// TIA Portal project "XSFW_TIA32801_A0" (V15.1) (continued)
REGION Network 14: Agrupa las fallas del proceso en una marca
   RUNG wire#powerrail
      I_Contact( "Fallas"."area de recorrido libre del pusher" )
      I_Contact( "Fallas"."caja trabada a la salida" )
      I_Contact( "Fallas".emergencia )
      I_Contact( "Fallas"."Falla de programación concatenadoras 1" )
      I_Contact( "Fallas"."Falla de programación concatenadoras 2" )
      I_Contact( "Fallas"."Falla de programación prioritarias 1" )
      I_Contact( "Fallas"."Falla de programación prioritarias 2" )
      I_Contact( "Fallas"."Falla en rele cadena" )
      I_Contact( "Fallas"."Falla en sensor de encolado" )
      I_Contact( "Fallas".falla_encoder )
      I_Contact( "Fallas".falla_sns_bsucc_ab )
      I_Contact( "Fallas".falla_sns_bsucc_ar )
      I_Contact( "Fallas"."Incrongruencia pusher" )
      I_Contact( "Fallas"."proteccion de torque" )
      I_Contact( "Fallas"."Falla en sensores del Pusher" )
      I_Contact( "Fallas"."Sensor pusher hacia adelante" )
      I_Contact( "Fallas"."Sin pegamento en el depósito" )
      I_Contact( "Fallas"."Falla de caja cerrada en cadena" )
      Coil( "Serie de fallas" )
   END_RUNG
   // the same network as SCL:
   "Serie de fallas" := NOT "Fallas"."area de recorrido libre del pusher" AND NOT "Fallas"."caja trabada a la salida" AND NOT "Fallas".emergencia AND NOT "Fallas"."Falla de programación concatenadoras 1" AND NOT "Fallas"."Falla de programación concatenadoras 2" AND NOT "Fallas"."Falla de programación prioritarias 1" AND NOT "Fallas"."Falla de programación prioritarias 2" AND NOT "Fallas"."Falla en rele cadena" AND NOT "Fallas"."Falla en sensor de encolado" AND NOT "Fallas".falla_encoder AND NOT "Fallas".falla_sns_bsucc_ab AND NOT "Fallas".falla_sns_bsucc_ar AND NOT "Fallas"."Incrongruencia pusher" AND NOT "Fallas"."proteccion de torque" AND NOT "Fallas"."Falla en sensores del Pusher" AND NOT "Fallas"."Sensor pusher hacia adelante" AND NOT "Fallas"."Sin pegamento en el depósito" AND NOT "Fallas"."Falla de caja cerrada en cadena";
END_REGION

REGION Network 15: Fallas en sensor atras del Pusher
   "Timer_DB7".TON(IN := "1s8" AND "oM_pusher" AND NOT "iSNSpush_atras", PT := T#350MS);
   "Fallas"."Falla en sensores del Pusher" := "Timer_DB7".Q;
END_REGION

REGION Network 16: Fallas en sensor adelante del Pusher
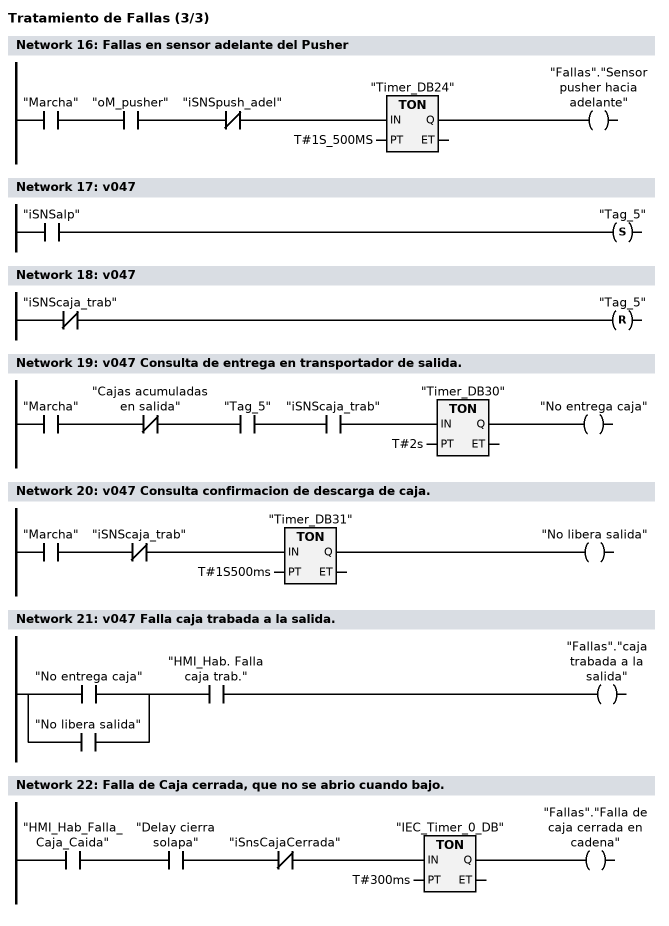
   "Timer_DB24".TON(IN := "Marcha" AND "oM_pusher" AND NOT "iSNSpush_adel", PT := T#1S_500MS);
   "Fallas"."Sensor pusher hacia adelante" := "Timer_DB24".Q;
END_REGION

REGION Network 17: v047
   RUNG wire#powerrail
      Contact( "iSNSalp" )
      S_Coil( "Tag_5" )
   END_RUNG
   // the same network as SCL:
   IF "iSNSalp" THEN "Tag_5" := TRUE; END_IF;
END_REGION

REGION Network 18: v047
   RUNG wire#powerrail
      I_Contact( "iSNScaja_trab" )
      R_Coil( "Tag_5" )
   END_RUNG
   // the same network as SCL:
   IF NOT "iSNScaja_trab" THEN "Tag_5" := FALSE; END_IF;
END_REGION

REGION Network 19: v047 Consulta de entrega en transportador de salida.
   "Timer_DB30".TON(IN := "Marcha" AND NOT "Cajas acumuladas en salida" AND "Tag_5" AND "iSNScaja_trab",
                    PT := T#2s);
   "No entrega caja" := "Timer_DB30".Q;
END_REGION

REGION Network 20: v047 Consulta confirmacion de descarga de caja.
   "Timer_DB31".TON(IN := "Marcha" AND NOT "iSNScaja_trab", PT := T#1S500ms);
   "No libera salida" := "Timer_DB31".Q;
END_REGION

REGION Network 21: v047 Falla caja trabada a la salida.
   RUNG wire#powerrail
      Contact( "No entrega caja" )
      wire#w1
      Contact( "HMI_Hab. Falla caja trab." )
      Coil( "Fallas"."caja trabada a la salida" )
   END_RUNG
   RUNG wire#powerrail
      Contact( "No libera salida" )
   END_RUNG wire#w1
   // the same network as SCL:
   "Fallas"."caja trabada a la salida" := ("No entrega caja" OR "No libera salida") AND "HMI_Hab. Falla caja trab.";
END_REGION

REGION Network 22: Falla de Caja cerrada, que no se abrio cuando bajo.
   "IEC_Timer_0_DB".TON(IN := "HMI_Hab_Falla_Caja_Caida" AND "Delay cierra solapa" AND NOT "iSnsCajaCerrada",
                        PT := T#300ms);
   "Fallas"."Falla de caja cerrada en cadena" := "IEC_Timer_0_DB".Q;
END_REGION
END_FUNCTION

FUNCTION "Salidas" : Void   // FC17, LAD
TITLE = Salidas del proceso (Modo Automático y Manual)
{ S7_Optimized_Access := 'TRUE' }
VERSION : 0.1
   VAR_TEMP   // added for the SCL form of the ladder/FBD networks
      _w1 : Bool;
   END_VAR
BEGIN

REGION Network 1: Activa la línea de emergencia del PLC
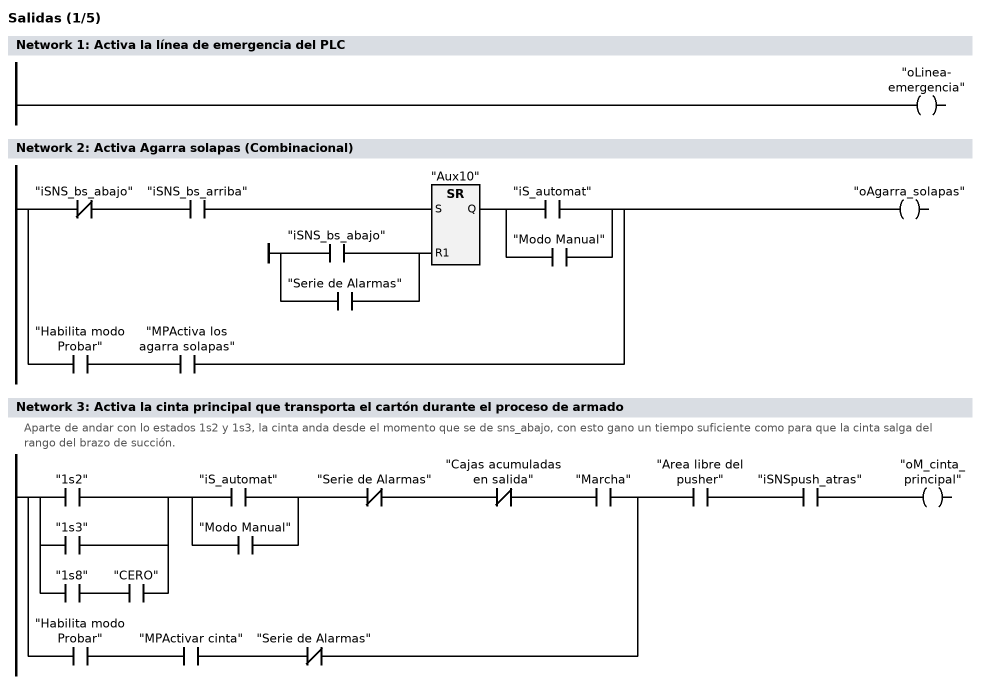
   RUNG wire#powerrail
      Coil( "oLinea-emergencia" )
   END_RUNG
   // the same network as SCL:
   "oLinea-emergencia" := TRUE;
END_REGION

REGION Network 2: Activa Agarra solapas (Combinacional)
   RUNG wire#powerrail
      I_Contact( "iSNS_bs_abajo" )
      Contact( "iSNS_bs_arriba" )
      S_SR(operand := "Aux10", r1 := wire#w1)
      wire#w2
      Contact( "iS_automat" )
      wire#w3
      Coil( "oAgarra_solapas" )
   END_RUNG
   RUNG wire#powerrail
      Contact( "iSNS_bs_abajo" )
   END_RUNG wire#w1
   RUNG wire#powerrail
      Contact( "Serie de Alarmas" )
   END_RUNG wire#w1
   RUNG wire#w2
      Contact( "Modo Manual" )
   END_RUNG wire#w3
   RUNG wire#powerrail
      Contact( "Habilita modo Probar" )
      Contact( "MPActiva los agarra solapas" )
   END_RUNG wire#w3
   // the same network as SCL:
   IF NOT "iSNS_bs_abajo" AND "iSNS_bs_arriba" THEN
       "Aux10" := TRUE;   // SR flip-flop
   END_IF;
   IF "iSNS_bs_abajo" OR "Serie de Alarmas" THEN "Aux10" := FALSE; END_IF;
   "oAgarra_solapas" := ("Aux10" AND ("iS_automat" OR "Modo Manual")) OR ("Habilita modo Probar" AND "MPActiva los agarra solapas");
END_REGION

REGION Network 3: Activa la cinta principal que transporta el cartón durante el proceso de armado
   // Aparte de andar con lo estados 1s2 y 1s3, la cinta anda desde el momento que se de sns_abajo, con esto gano un tiempo suficiente como para que la cinta salga del rango del brazo de succión.
   RUNG wire#powerrail
      Contact( "1s2" )
      wire#w1
      Contact( "iS_automat" )
      wire#w2
      I_Contact( "Serie de Alarmas" )
      I_Contact( "Cajas acumuladas en salida" )
      Contact( "Marcha" )
      wire#w3
      Contact( "Area libre del pusher" )
      Contact( "iSNSpush_atras" )
      Coil( "oM_cinta_principal" )
   END_RUNG
   RUNG wire#powerrail
      Contact( "1s3" )
   END_RUNG wire#w1
   RUNG wire#powerrail
      Contact( "1s8" )
      Contact( "CERO" )
   END_RUNG wire#w1
   RUNG wire#w1
      Contact( "Modo Manual" )
   END_RUNG wire#w2
   RUNG wire#powerrail
      Contact( "Habilita modo Probar" )
      Contact( "MPActivar cinta" )
      I_Contact( "Serie de Alarmas" )
   END_RUNG wire#w3
   // the same network as SCL:
   "oM_cinta_principal" := ((("1s2" OR "1s3" OR ("1s8" AND "CERO")) AND ("iS_automat" OR "Modo Manual") AND NOT "Serie de Alarmas" AND NOT "Cajas acumuladas en salida" AND "Marcha") OR ("Habilita modo Probar" AND "MPActivar cinta" AND NOT "Serie de Alarmas")) AND "Area libre del pusher" AND "iSNSpush_atras";
END_REGION

REGION Network 4: Activa la boquilla encoladora.
   // Activa la boquilla encoladora a partir de determinados valores del encoder.El sensor de área de encolado se utiliza para fines de seguridad. El inicio de encolado se valida con la marca "aux encol 2"
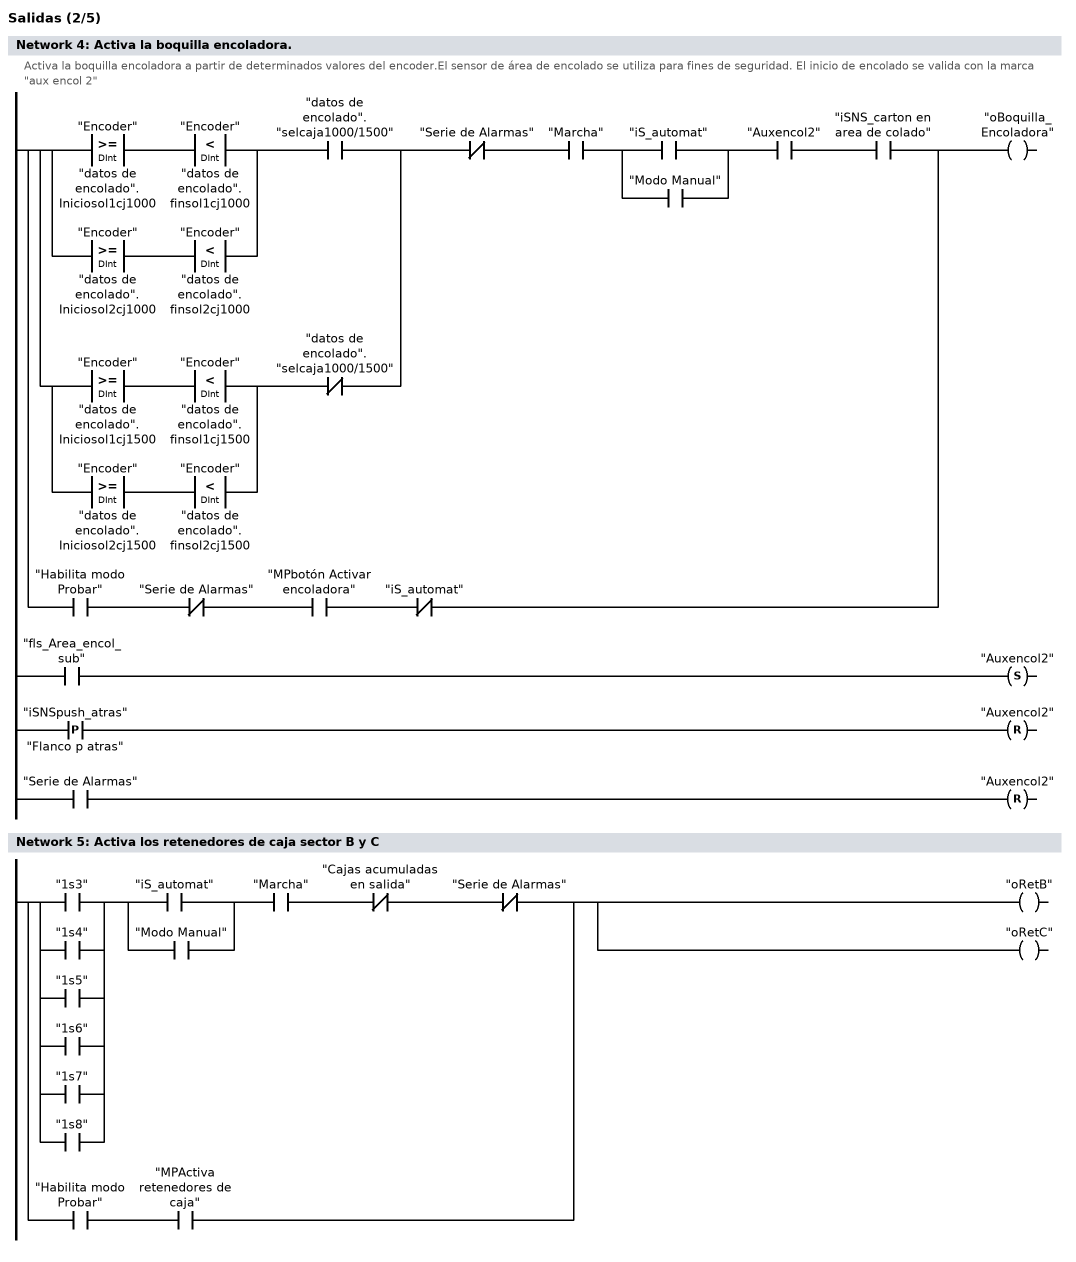
   RUNG wire#powerrail
      { S7_Templates := "SrcType := DInt" } GE_Contact(in1 := "Encoder", in2 := "datos de encolado".Iniciosol1cj1000)
      { S7_Templates := "SrcType := DInt" } LT_Contact(in1 := "Encoder", in2 := "datos de encolado".finsol1cj1000)
      wire#w1
      Contact( "datos de encolado"."selcaja1000/1500" )
      wire#w2
      I_Contact( "Serie de Alarmas" )
      Contact( "Marcha" )
      wire#w4
      Contact( "iS_automat" )
      wire#w5
      Contact( "Auxencol2" )
      Contact( "iSNS_carton en area de colado" )
      wire#w6
      Coil( "oBoquilla_Encoladora" )
   END_RUNG
   RUNG wire#powerrail
      { S7_Templates := "SrcType := DInt" } GE_Contact(in1 := "Encoder", in2 := "datos de encolado".Iniciosol2cj1000)
      { S7_Templates := "SrcType := DInt" } LT_Contact(in1 := "Encoder", in2 := "datos de encolado".finsol2cj1000)
   END_RUNG wire#w1
   RUNG wire#powerrail
      { S7_Templates := "SrcType := DInt" } GE_Contact(in1 := "Encoder", in2 := "datos de encolado".Iniciosol1cj1500)
      { S7_Templates := "SrcType := DInt" } LT_Contact(in1 := "Encoder", in2 := "datos de encolado".finsol1cj1500)
      wire#w3
      I_Contact( "datos de encolado"."selcaja1000/1500" )
   END_RUNG wire#w2
   RUNG wire#powerrail
      { S7_Templates := "SrcType := DInt" } GE_Contact(in1 := "Encoder", in2 := "datos de encolado".Iniciosol2cj1500)
      { S7_Templates := "SrcType := DInt" } LT_Contact(in1 := "Encoder", in2 := "datos de encolado".finsol2cj1500)
   END_RUNG wire#w3
   RUNG wire#w4
      Contact( "Modo Manual" )
   END_RUNG wire#w5
   RUNG wire#powerrail
      Contact( "Habilita modo Probar" )
      I_Contact( "Serie de Alarmas" )
      Contact( "MPbotón Activar encoladora" )
      I_Contact( "iS_automat" )
   END_RUNG wire#w6
   RUNG wire#powerrail
      Contact( "fls_Area_encol_sub" )
      S_Coil( "Auxencol2" )
   END_RUNG
   RUNG wire#powerrail
      P_Contact(operand := "iSNSpush_atras", bit := "Flanco p atras")
      R_Coil( "Auxencol2" )
   END_RUNG
   RUNG wire#powerrail
      Contact( "Serie de Alarmas" )
      R_Coil( "Auxencol2" )
   END_RUNG
   // the same network as SCL:
   "oBoquilla_Encoladora" := (((((("Encoder" >= "datos de encolado".Iniciosol1cj1000) AND ("Encoder" < "datos de encolado".finsol1cj1000)) OR (("Encoder" >= "datos de encolado".Iniciosol2cj1000) AND ("Encoder" < "datos de encolado".finsol2cj1000))) AND "datos de encolado"."selcaja1000/1500") OR (((("Encoder" >= "datos de encolado".Iniciosol1cj1500) AND ("Encoder" < "datos de encolado".finsol1cj1500)) OR (("Encoder" >= "datos de encolado".Iniciosol2cj1500) AND ("Encoder" < "datos de encolado".finsol2cj1500))) AND NOT "datos de encolado"."selcaja1000/1500")) AND NOT "Serie de Alarmas" AND "Marcha" AND ("iS_automat" OR "Modo Manual") AND "Auxencol2" AND "iSNS_carton en area de colado") OR ("Habilita modo Probar" AND NOT "Serie de Alarmas" AND "MPbotón Activar encoladora" AND NOT "iS_automat");
   IF "fls_Area_encol_sub" THEN "Auxencol2" := TRUE; END_IF;
   #_w1 := "iSNSpush_atras" AND NOT "Flanco p atras";   // rising edge of "iSNSpush_atras"
   "Flanco p atras" := "iSNSpush_atras";
   IF #_w1 THEN "Auxencol2" := FALSE; END_IF;
   IF "Serie de Alarmas" THEN "Auxencol2" := FALSE; END_IF;
END_REGION

REGION Network 5: Activa los retenedores de caja sector B y C
   RUNG wire#powerrail
      Contact( "1s3" )
      wire#w1
      Contact( "iS_automat" )
      wire#w2
      Contact( "Marcha" )
      I_Contact( "Cajas acumuladas en salida" )
      I_Contact( "Serie de Alarmas" )
      wire#w3
      Coil( "oRetB" )
   END_RUNG
   RUNG wire#powerrail
      Contact( "1s4" )
   END_RUNG wire#w1
   RUNG wire#powerrail
      Contact( "1s5" )
   END_RUNG wire#w1
   RUNG wire#powerrail
      Contact( "1s6" )
   END_RUNG wire#w1
   RUNG wire#powerrail
      Contact( "1s7" )
   END_RUNG wire#w1
   RUNG wire#powerrail
      Contact( "1s8" )
   END_RUNG wire#w1
   RUNG wire#w1
      Contact( "Modo Manual" )
   END_RUNG wire#w2
   RUNG wire#powerrail
      Contact( "Habilita modo Probar" )
      Contact( "MPActiva retenedores de caja" )
   END_RUNG wire#w3
   RUNG wire#w3
      Coil( "oRetC" )
   END_RUNG
   // the same network as SCL:
   "oRetB" := (("1s3" OR "1s4" OR "1s5" OR "1s6" OR "1s7" OR "1s8") AND ("iS_automat" OR "Modo Manual") AND "Marcha" AND NOT "Cajas acumuladas en salida" AND NOT "Serie de Alarmas") OR ("Habilita modo Probar" AND "MPActiva retenedores de caja");
   "oRetC" := "oRetB";
END_REGION

REGION Network 6
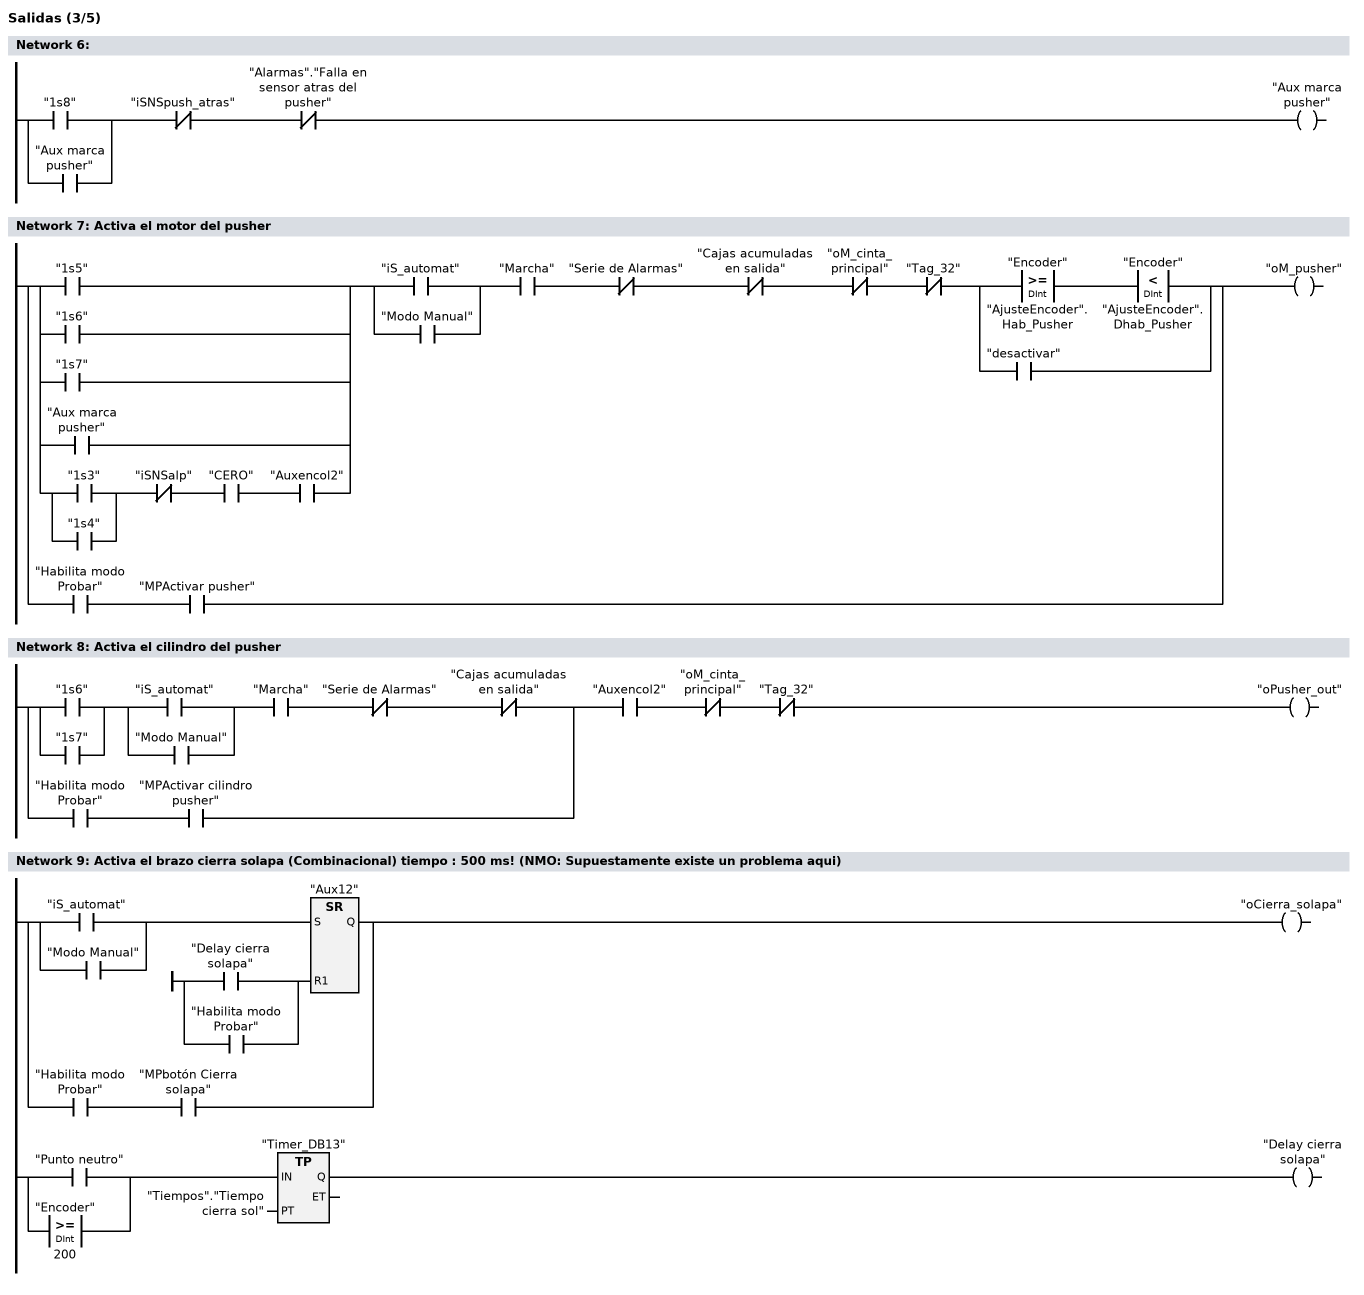
   RUNG wire#powerrail
      Contact( "1s8" )
      wire#w1
      I_Contact( "iSNSpush_atras" )
      I_Contact( "Alarmas"."Falla en sensor atras del pusher" )
      Coil( "Aux marca pusher" )
   END_RUNG
   RUNG wire#powerrail
      Contact( "Aux marca pusher" )
   END_RUNG wire#w1
   // the same network as SCL:
   "Aux marca pusher" := ("1s8" OR "Aux marca pusher") AND NOT "iSNSpush_atras" AND NOT "Alarmas"."Falla en sensor atras del pusher";
END_REGION

REGION Network 7: Activa el motor del pusher
   RUNG wire#powerrail
      Contact( "1s5" )
      wire#w1
      Contact( "iS_automat" )
      wire#w3
      Contact( "Marcha" )
      I_Contact( "Serie de Alarmas" )
      I_Contact( "Cajas acumuladas en salida" )
      I_Contact( "oM_cinta_principal" )
      I_Contact( "Tag_32" )
      wire#w4
      { S7_Templates := "SrcType := DInt" } GE_Contact(in1 := "Encoder", in2 := "AjusteEncoder".Hab_Pusher)
      { S7_Templates := "SrcType := DInt" } LT_Contact(in1 := "Encoder", in2 := "AjusteEncoder".Dhab_Pusher)
      wire#w5
      Coil( "oM_pusher" )
   END_RUNG
   RUNG wire#powerrail
      Contact( "1s6" )
   END_RUNG wire#w1
   RUNG wire#powerrail
      Contact( "1s7" )
   END_RUNG wire#w1
   RUNG wire#powerrail
      Contact( "Aux marca pusher" )
   END_RUNG wire#w1
   RUNG wire#powerrail
      Contact( "1s3" )
      wire#w2
      I_Contact( "iSNSalp" )
      Contact( "CERO" )
      Contact( "Auxencol2" )
   END_RUNG wire#w1
   RUNG wire#powerrail
      Contact( "1s4" )
   END_RUNG wire#w2
   RUNG wire#w1
      Contact( "Modo Manual" )
   END_RUNG wire#w3
   RUNG wire#w4
      Contact( "desactivar" )
   END_RUNG wire#w5
   RUNG wire#powerrail
      Contact( "Habilita modo Probar" )
      Contact( "MPActivar pusher" )
   END_RUNG wire#w5
   // the same network as SCL:
   "oM_pusher" := (("1s5" OR "1s6" OR "1s7" OR "Aux marca pusher" OR (("1s3" OR "1s4") AND NOT "iSNSalp" AND "CERO" AND "Auxencol2")) AND ("iS_automat" OR "Modo Manual") AND "Marcha" AND NOT "Serie de Alarmas" AND NOT "Cajas acumuladas en salida" AND NOT "oM_cinta_principal" AND NOT "Tag_32" AND ((("Encoder" >= "AjusteEncoder".Hab_Pusher) AND ("Encoder" < "AjusteEncoder".Dhab_Pusher)) OR "desactivar")) OR ("Habilita modo Probar" AND "MPActivar pusher");
END_REGION

REGION Network 8: Activa el cilindro del pusher
   RUNG wire#powerrail
      Contact( "1s6" )
      wire#w1
      Contact( "iS_automat" )
      wire#w2
      Contact( "Marcha" )
      I_Contact( "Serie de Alarmas" )
      I_Contact( "Cajas acumuladas en salida" )
      wire#w3
      Contact( "Auxencol2" )
      I_Contact( "oM_cinta_principal" )
      I_Contact( "Tag_32" )
      Coil( "oPusher_out" )
   END_RUNG
   RUNG wire#powerrail
      Contact( "1s7" )
   END_RUNG wire#w1
   RUNG wire#w1
      Contact( "Modo Manual" )
   END_RUNG wire#w2
   RUNG wire#powerrail
      Contact( "Habilita modo Probar" )
      Contact( "MPActivar cilindro pusher" )
   END_RUNG wire#w3
   // the same network as SCL:
   "oPusher_out" := ((("1s6" OR "1s7") AND ("iS_automat" OR "Modo Manual") AND "Marcha" AND NOT "Serie de Alarmas" AND NOT "Cajas acumuladas en salida") OR ("Habilita modo Probar" AND "MPActivar cilindro pusher")) AND "Auxencol2" AND NOT "oM_cinta_principal" AND NOT "Tag_32";
END_REGION

REGION Network 9: Activa el brazo cierra solapa (Combinacional) tiempo : 500 ms! (NMO: Supuestamente existe un problema aqui)
   IF "iS_automat" OR "Modo Manual" THEN
       "Aux12" := TRUE;   // SR flip-flop
   END_IF;
   IF "Delay cierra solapa" OR "Habilita modo Probar" THEN "Aux12" := FALSE; END_IF;
   "oCierra_solapa" := "Aux12" OR ("Habilita modo Probar" AND "MPbotón Cierra solapa");
   "Timer_DB13".TP(IN := "Punto neutro" OR ("Encoder" >= 200), PT := "Tiempos"."Tiempo cierra sol");
   "Delay cierra solapa" := "Timer_DB13".Q;
END_REGION

REGION Network 10: Activa la pinza sssssss
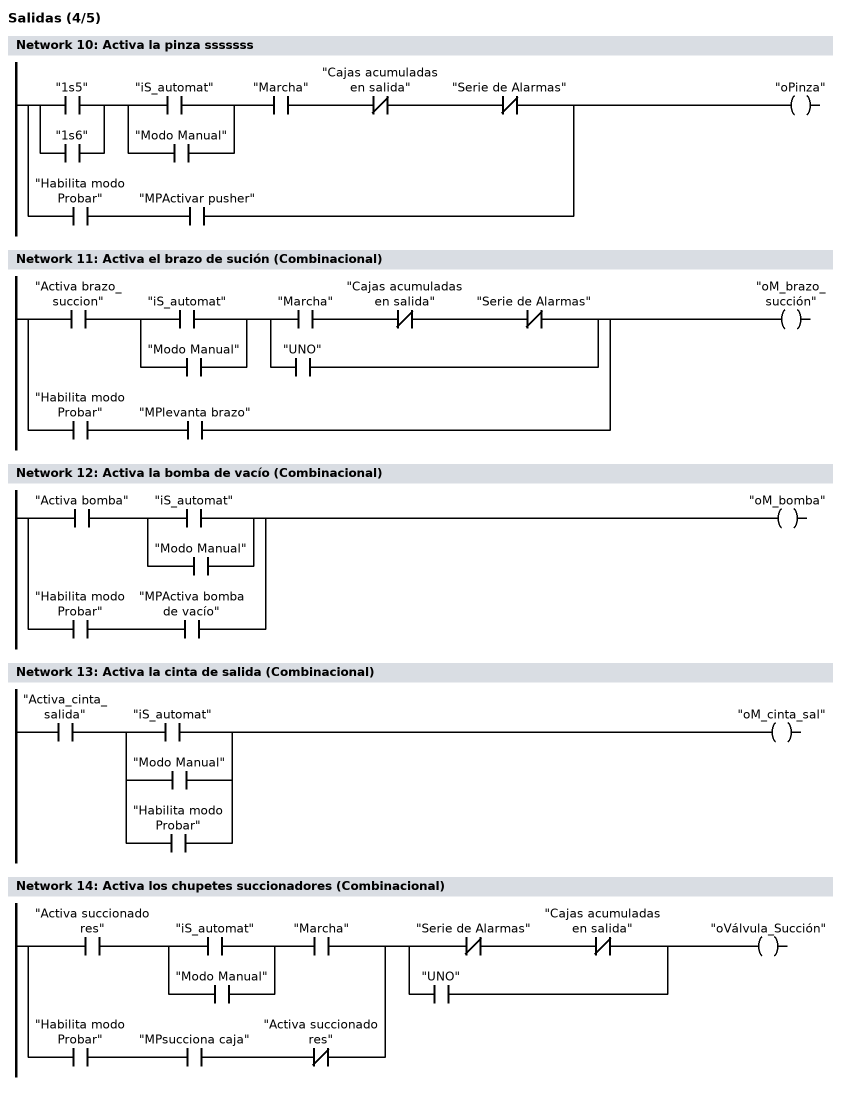
   RUNG wire#powerrail
      Contact( "1s5" )
      wire#w1
      Contact( "iS_automat" )
      wire#w2
      Contact( "Marcha" )
      I_Contact( "Cajas acumuladas en salida" )
      I_Contact( "Serie de Alarmas" )
      wire#w3
      Coil( "oPinza" )
   END_RUNG
   RUNG wire#powerrail
      Contact( "1s6" )
   END_RUNG wire#w1
   RUNG wire#w1
      Contact( "Modo Manual" )
   END_RUNG wire#w2
   RUNG wire#powerrail
      Contact( "Habilita modo Probar" )
      Contact( "MPActivar pusher" )
   END_RUNG wire#w3
   // the same network as SCL:
   "oPinza" := (("1s5" OR "1s6") AND ("iS_automat" OR "Modo Manual") AND "Marcha" AND NOT "Cajas acumuladas en salida" AND NOT "Serie de Alarmas") OR ("Habilita modo Probar" AND "MPActivar pusher");
END_REGION

REGION Network 11: Activa el brazo de sución (Combinacional)
   RUNG wire#powerrail
      Contact( "Activa brazo_succion" )
      wire#w1
      Contact( "iS_automat" )
      wire#w2
      Contact( "Marcha" )
      I_Contact( "Cajas acumuladas en salida" )
      I_Contact( "Serie de Alarmas" )
      wire#w3
      Coil( "oM_brazo_succión" )
   END_RUNG
   RUNG wire#w1
      Contact( "Modo Manual" )
   END_RUNG wire#w2
   RUNG wire#w2
      Contact( "UNO" )
   END_RUNG wire#w3
   RUNG wire#powerrail
      Contact( "Habilita modo Probar" )
      Contact( "MPlevanta brazo" )
   END_RUNG wire#w3
   // the same network as SCL:
   "oM_brazo_succión" := ("Activa brazo_succion" AND ("iS_automat" OR "Modo Manual") AND (("Marcha" AND NOT "Cajas acumuladas en salida" AND NOT "Serie de Alarmas") OR "UNO")) OR ("Habilita modo Probar" AND "MPlevanta brazo");
END_REGION

REGION Network 12: Activa la bomba de vacío (Combinacional)
   RUNG wire#powerrail
      Contact( "Activa bomba" )
      wire#w1
      Contact( "iS_automat" )
      wire#w2
      Coil( "oM_bomba" )
   END_RUNG
   RUNG wire#w1
      Contact( "Modo Manual" )
   END_RUNG wire#w2
   RUNG wire#powerrail
      Contact( "Habilita modo Probar" )
      Contact( "MPActiva bomba de vacío" )
   END_RUNG wire#w2
   // the same network as SCL:
   "oM_bomba" := ("Activa bomba" AND ("iS_automat" OR "Modo Manual")) OR ("Habilita modo Probar" AND "MPActiva bomba de vacío");
END_REGION

REGION Network 13: Activa la cinta de salida (Combinacional)
   RUNG wire#powerrail
      Contact( "Activa_cinta_salida" )
      wire#w1
      Contact( "iS_automat" )
      wire#w2
      Coil( "oM_cinta_sal" )
   END_RUNG
   RUNG wire#w1
      Contact( "Modo Manual" )
   END_RUNG wire#w2
   RUNG wire#w1
      Contact( "Habilita modo Probar" )
   END_RUNG wire#w2
   // the same network as SCL:
   "oM_cinta_sal" := "Activa_cinta_salida" AND ("iS_automat" OR "Modo Manual" OR "Habilita modo Probar");
END_REGION

REGION Network 14: Activa los chupetes succionadores (Combinacional)
   RUNG wire#powerrail
      Contact( "Activa succionadores" )
      wire#w1
      Contact( "iS_automat" )
      wire#w2
      Contact( "Marcha" )
      wire#w3
      I_Contact( "Serie de Alarmas" )
      I_Contact( "Cajas acumuladas en salida" )
      wire#w4
      Coil( "oVálvula_Succión" )
   END_RUNG
   RUNG wire#w1
      Contact( "Modo Manual" )
   END_RUNG wire#w2
   RUNG wire#powerrail
      Contact( "Habilita modo Probar" )
      Contact( "MPsucciona caja" )
      I_Contact( "Activa succionadores" )
   END_RUNG wire#w3
   RUNG wire#w3
      Contact( "UNO" )
   END_RUNG wire#w4
   // the same network as SCL:
   "oVálvula_Succión" := (("Activa succionadores" AND ("iS_automat" OR "Modo Manual") AND "Marcha") OR ("Habilita modo Probar" AND "MPsucciona caja" AND NOT "Activa succionadores")) AND ((NOT "Serie de Alarmas" AND NOT "Cajas acumuladas en salida") OR "UNO");
END_REGION

REGION Network 15: Pone en marcha la armadora (la entrada EXT no existe , tampoco la "opacker" )
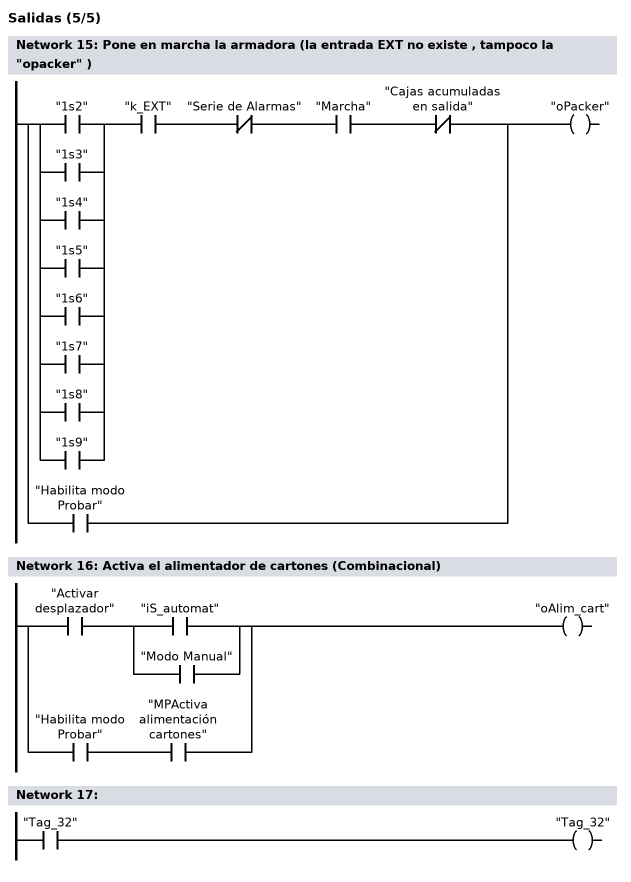
   RUNG wire#powerrail
      Contact( "1s2" )
      wire#w1
      Contact( "k_EXT" )
      I_Contact( "Serie de Alarmas" )
      Contact( "Marcha" )
      I_Contact( "Cajas acumuladas en salida" )
      wire#w2
      Coil( "oPacker" )
   END_RUNG
   RUNG wire#powerrail
      Contact( "1s3" )
   END_RUNG wire#w1
   RUNG wire#powerrail
      Contact( "1s4" )
   END_RUNG wire#w1
   RUNG wire#powerrail
      Contact( "1s5" )
   END_RUNG wire#w1
   RUNG wire#powerrail
      Contact( "1s6" )
   END_RUNG wire#w1
   RUNG wire#powerrail
      Contact( "1s7" )
   END_RUNG wire#w1
   RUNG wire#powerrail
      Contact( "1s8" )
   END_RUNG wire#w1
   RUNG wire#powerrail
      Contact( "1s9" )
   END_RUNG wire#w1
   RUNG wire#powerrail
      Contact( "Habilita modo Probar" )
   END_RUNG wire#w2
   // the same network as SCL:
   "oPacker" := (("1s2" OR "1s3" OR "1s4" OR "1s5" OR "1s6" OR "1s7" OR "1s8" OR "1s9") AND "k_EXT" AND NOT "Serie de Alarmas" AND "Marcha" AND NOT "Cajas acumuladas en salida") OR "Habilita modo Probar";
END_REGION

REGION Network 16: Activa el alimentador de cartones (Combinacional)
   RUNG wire#powerrail
      Contact( "Activar desplazador" )
      wire#w1
      Contact( "iS_automat" )
      wire#w2
      Coil( "oAlim_cart" )
   END_RUNG
   RUNG wire#w1
      Contact( "Modo Manual" )
   END_RUNG wire#w2
   RUNG wire#powerrail
      Contact( "Habilita modo Probar" )
      Contact( "MPActiva alimentación cartones" )
   END_RUNG wire#w2
   // the same network as SCL:
   "oAlim_cart" := ("Activar desplazador" AND ("iS_automat" OR "Modo Manual")) OR ("Habilita modo Probar" AND "MPActiva alimentación cartones");
END_REGION

REGION Network 17
   RUNG wire#powerrail
      Contact( "Tag_32" )
      Coil( "Tag_32" )
   END_RUNG
   // the same network as SCL:
   "Tag_32" := "Tag_32";
END_REGION
END_FUNCTION

FUNCTION "MAQ-EST-32-SEC1" : Void   // FC18, LAD
{ S7_Optimized_Access := 'TRUE' }
VERSION : 0.1
   VAR_INPUT
      Concatenadora : DWord;
      Prioritaria : DWord;
   END_VAR
   VAR_IN_OUT
      "Falla Prioritarias" : Bool;
      "Error Concatenadoras" : Bool;
      Estado : DWord;
   END_VAR
BEGIN

REGION Network 1: Falla Prioritarias
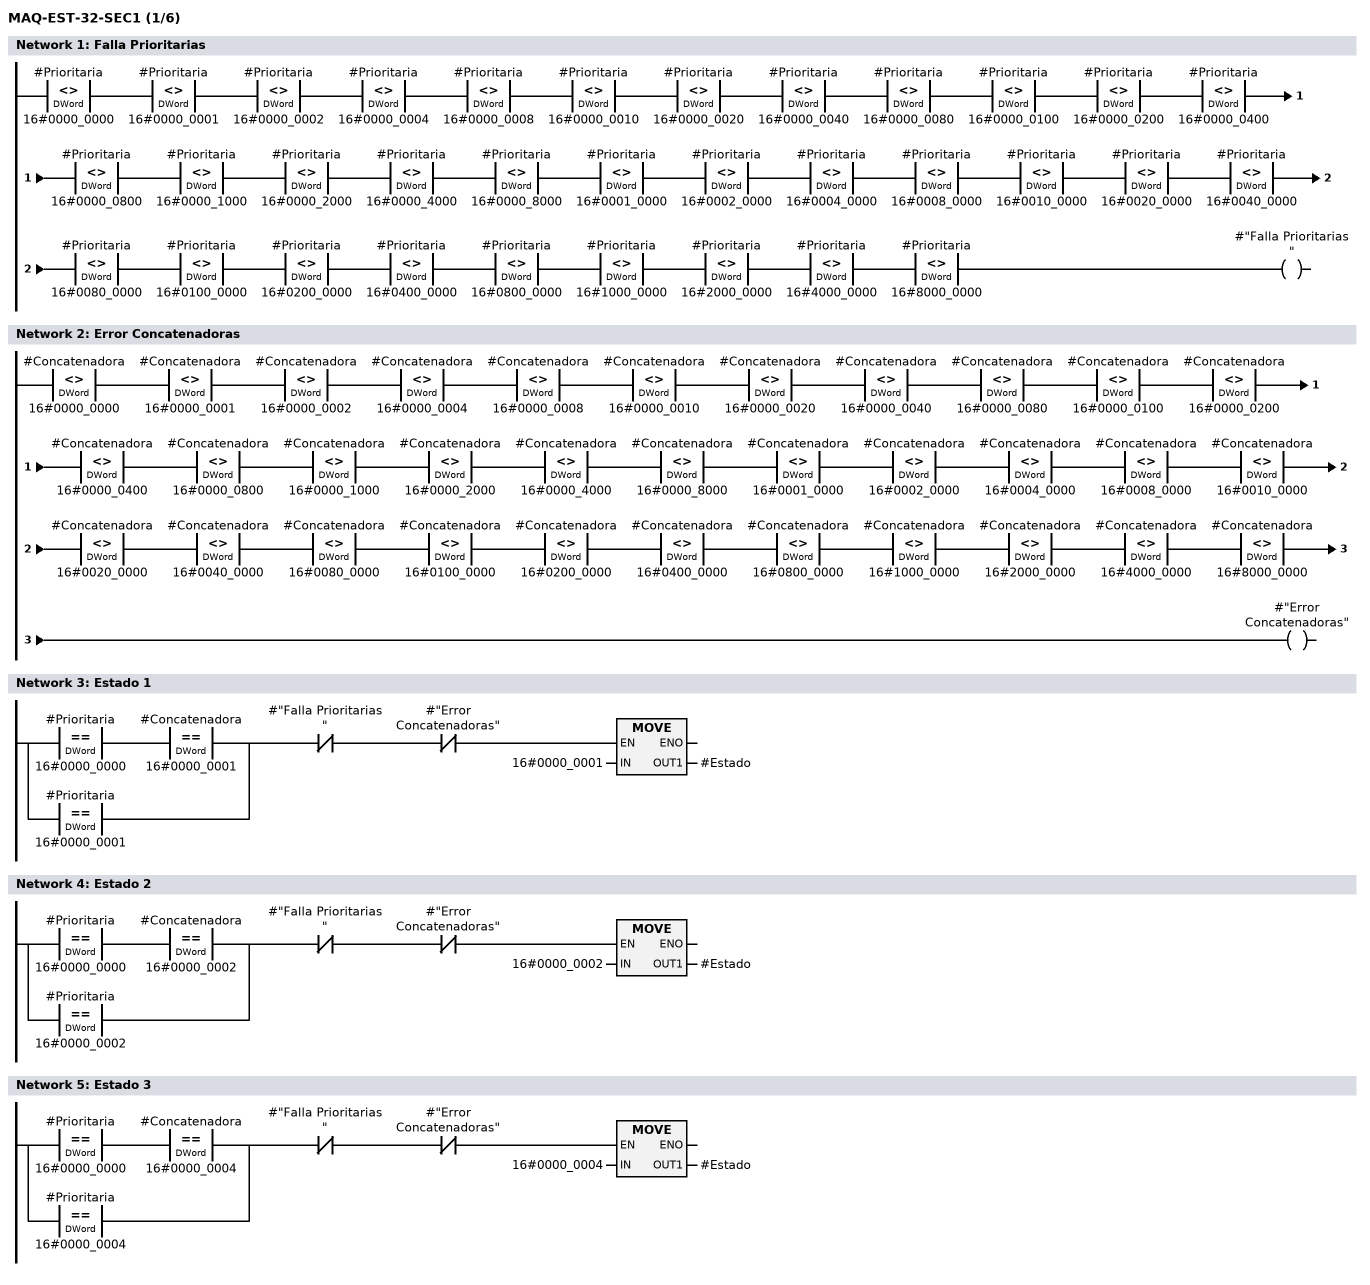
   RUNG wire#powerrail
      { S7_Templates := "SrcType := DWord" } NE_Contact(in1 := #Prioritaria, in2 := 16#0000_0000)
      { S7_Templates := "SrcType := DWord" } NE_Contact(in1 := #Prioritaria, in2 := 16#0000_0001)
      { S7_Templates := "SrcType := DWord" } NE_Contact(in1 := #Prioritaria, in2 := 16#0000_0002)
      { S7_Templates := "SrcType := DWord" } NE_Contact(in1 := #Prioritaria, in2 := 16#0000_0004)
      { S7_Templates := "SrcType := DWord" } NE_Contact(in1 := #Prioritaria, in2 := 16#0000_0008)
      { S7_Templates := "SrcType := DWord" } NE_Contact(in1 := #Prioritaria, in2 := 16#0000_0010)
      { S7_Templates := "SrcType := DWord" } NE_Contact(in1 := #Prioritaria, in2 := 16#0000_0020)
      { S7_Templates := "SrcType := DWord" } NE_Contact(in1 := #Prioritaria, in2 := 16#0000_0040)
      { S7_Templates := "SrcType := DWord" } NE_Contact(in1 := #Prioritaria, in2 := 16#0000_0080)
      { S7_Templates := "SrcType := DWord" } NE_Contact(in1 := #Prioritaria, in2 := 16#0000_0100)
      { S7_Templates := "SrcType := DWord" } NE_Contact(in1 := #Prioritaria, in2 := 16#0000_0200)
      { S7_Templates := "SrcType := DWord" } NE_Contact(in1 := #Prioritaria, in2 := 16#0000_0400)
      { S7_Templates := "SrcType := DWord" } NE_Contact(in1 := #Prioritaria, in2 := 16#0000_0800)
      { S7_Templates := "SrcType := DWord" } NE_Contact(in1 := #Prioritaria, in2 := 16#0000_1000)
      { S7_Templates := "SrcType := DWord" } NE_Contact(in1 := #Prioritaria, in2 := 16#0000_2000)
      { S7_Templates := "SrcType := DWord" } NE_Contact(in1 := #Prioritaria, in2 := 16#0000_4000)
      { S7_Templates := "SrcType := DWord" } NE_Contact(in1 := #Prioritaria, in2 := 16#0000_8000)
      { S7_Templates := "SrcType := DWord" } NE_Contact(in1 := #Prioritaria, in2 := 16#0001_0000)
      { S7_Templates := "SrcType := DWord" } NE_Contact(in1 := #Prioritaria, in2 := 16#0002_0000)
      { S7_Templates := "SrcType := DWord" } NE_Contact(in1 := #Prioritaria, in2 := 16#0004_0000)
      { S7_Templates := "SrcType := DWord" } NE_Contact(in1 := #Prioritaria, in2 := 16#0008_0000)
      { S7_Templates := "SrcType := DWord" } NE_Contact(in1 := #Prioritaria, in2 := 16#0010_0000)
      { S7_Templates := "SrcType := DWord" } NE_Contact(in1 := #Prioritaria, in2 := 16#0020_0000)
      { S7_Templates := "SrcType := DWord" } NE_Contact(in1 := #Prioritaria, in2 := 16#0040_0000)
      { S7_Templates := "SrcType := DWord" } NE_Contact(in1 := #Prioritaria, in2 := 16#0080_0000)
      { S7_Templates := "SrcType := DWord" } NE_Contact(in1 := #Prioritaria, in2 := 16#0100_0000)
      { S7_Templates := "SrcType := DWord" } NE_Contact(in1 := #Prioritaria, in2 := 16#0200_0000)
      { S7_Templates := "SrcType := DWord" } NE_Contact(in1 := #Prioritaria, in2 := 16#0400_0000)
      { S7_Templates := "SrcType := DWord" } NE_Contact(in1 := #Prioritaria, in2 := 16#0800_0000)
      { S7_Templates := "SrcType := DWord" } NE_Contact(in1 := #Prioritaria, in2 := 16#1000_0000)
      { S7_Templates := "SrcType := DWord" } NE_Contact(in1 := #Prioritaria, in2 := 16#2000_0000)
      { S7_Templates := "SrcType := DWord" } NE_Contact(in1 := #Prioritaria, in2 := 16#4000_0000)
      { S7_Templates := "SrcType := DWord" } NE_Contact(in1 := #Prioritaria, in2 := 16#8000_0000)
      Coil( #"Falla Prioritarias" )
   END_RUNG
   // the same network as SCL:
   #"Falla Prioritarias" := (#Prioritaria <> 16#0000_0000) AND (#Prioritaria <> 16#0000_0001) AND (#Prioritaria <> 16#0000_0002) AND (#Prioritaria <> 16#0000_0004) AND (#Prioritaria <> 16#0000_0008) AND (#Prioritaria <> 16#0000_0010) AND (#Prioritaria <> 16#0000_0020) AND (#Prioritaria <> 16#0000_0040) AND (#Prioritaria <> 16#0000_0080) AND (#Prioritaria <> 16#0000_0100) AND (#Prioritaria <> 16#0000_0200) AND (#Prioritaria <> 16#0000_0400) AND (#Prioritaria <> 16#0000_0800) AND (#Prioritaria <> 16#0000_1000) AND (#Prioritaria <> 16#0000_2000) AND (#Prioritaria <> 16#0000_4000) AND (#Prioritaria <> 16#0000_8000) AND (#Prioritaria <> 16#0001_0000) AND (#Prioritaria <> 16#0002_0000) AND (#Prioritaria <> 16#0004_0000) AND (#Prioritaria <> 16#0008_0000) AND (#Prioritaria <> 16#0010_0000) AND (#Prioritaria <> 16#0020_0000) AND (#Prioritaria <> 16#0040_0000) AND (#Prioritaria <> 16#0080_0000) AND (#Prioritaria <> 16#0100_0000) AND (#Prioritaria <> 16#0200_0000) AND (#Prioritaria <> 16#0400_0000) AND (#Prioritaria <> 16#0800_0000) AND (#Prioritaria <> 16#1000_0000) AND (#Prioritaria <> 16#2000_0000) AND (#Prioritaria <> 16#4000_0000) AND (#Prioritaria <> 16#8000_0000);
END_REGION

REGION Network 2: Error Concatenadoras
   RUNG wire#powerrail
      { S7_Templates := "SrcType := DWord" } NE_Contact(in1 := #Concatenadora, in2 := 16#0000_0000)
      { S7_Templates := "SrcType := DWord" } NE_Contact(in1 := #Concatenadora, in2 := 16#0000_0001)
      { S7_Templates := "SrcType := DWord" } NE_Contact(in1 := #Concatenadora, in2 := 16#0000_0002)
      { S7_Templates := "SrcType := DWord" } NE_Contact(in1 := #Concatenadora, in2 := 16#0000_0004)
      { S7_Templates := "SrcType := DWord" } NE_Contact(in1 := #Concatenadora, in2 := 16#0000_0008)
      { S7_Templates := "SrcType := DWord" } NE_Contact(in1 := #Concatenadora, in2 := 16#0000_0010)
      { S7_Templates := "SrcType := DWord" } NE_Contact(in1 := #Concatenadora, in2 := 16#0000_0020)
      { S7_Templates := "SrcType := DWord" } NE_Contact(in1 := #Concatenadora, in2 := 16#0000_0040)
      { S7_Templates := "SrcType := DWord" } NE_Contact(in1 := #Concatenadora, in2 := 16#0000_0080)
      { S7_Templates := "SrcType := DWord" } NE_Contact(in1 := #Concatenadora, in2 := 16#0000_0100)
      { S7_Templates := "SrcType := DWord" } NE_Contact(in1 := #Concatenadora, in2 := 16#0000_0200)
      { S7_Templates := "SrcType := DWord" } NE_Contact(in1 := #Concatenadora, in2 := 16#0000_0400)
      { S7_Templates := "SrcType := DWord" } NE_Contact(in1 := #Concatenadora, in2 := 16#0000_0800)
      { S7_Templates := "SrcType := DWord" } NE_Contact(in1 := #Concatenadora, in2 := 16#0000_1000)
      { S7_Templates := "SrcType := DWord" } NE_Contact(in1 := #Concatenadora, in2 := 16#0000_2000)
      { S7_Templates := "SrcType := DWord" } NE_Contact(in1 := #Concatenadora, in2 := 16#0000_4000)
      { S7_Templates := "SrcType := DWord" } NE_Contact(in1 := #Concatenadora, in2 := 16#0000_8000)
      { S7_Templates := "SrcType := DWord" } NE_Contact(in1 := #Concatenadora, in2 := 16#0001_0000)
      { S7_Templates := "SrcType := DWord" } NE_Contact(in1 := #Concatenadora, in2 := 16#0002_0000)
      { S7_Templates := "SrcType := DWord" } NE_Contact(in1 := #Concatenadora, in2 := 16#0004_0000)
      { S7_Templates := "SrcType := DWord" } NE_Contact(in1 := #Concatenadora, in2 := 16#0008_0000)
      { S7_Templates := "SrcType := DWord" } NE_Contact(in1 := #Concatenadora, in2 := 16#0010_0000)
      { S7_Templates := "SrcType := DWord" } NE_Contact(in1 := #Concatenadora, in2 := 16#0020_0000)
      { S7_Templates := "SrcType := DWord" } NE_Contact(in1 := #Concatenadora, in2 := 16#0040_0000)
      { S7_Templates := "SrcType := DWord" } NE_Contact(in1 := #Concatenadora, in2 := 16#0080_0000)
      { S7_Templates := "SrcType := DWord" } NE_Contact(in1 := #Concatenadora, in2 := 16#0100_0000)
      { S7_Templates := "SrcType := DWord" } NE_Contact(in1 := #Concatenadora, in2 := 16#0200_0000)
      { S7_Templates := "SrcType := DWord" } NE_Contact(in1 := #Concatenadora, in2 := 16#0400_0000)
      { S7_Templates := "SrcType := DWord" } NE_Contact(in1 := #Concatenadora, in2 := 16#0800_0000)
      { S7_Templates := "SrcType := DWord" } NE_Contact(in1 := #Concatenadora, in2 := 16#1000_0000)
      { S7_Templates := "SrcType := DWord" } NE_Contact(in1 := #Concatenadora, in2 := 16#2000_0000)
      { S7_Templates := "SrcType := DWord" } NE_Contact(in1 := #Concatenadora, in2 := 16#4000_0000)
      { S7_Templates := "SrcType := DWord" } NE_Contact(in1 := #Concatenadora, in2 := 16#8000_0000)
      Coil( #"Error Concatenadoras" )
   END_RUNG
   // the same network as SCL:
   #"Error Concatenadoras" := (#Concatenadora <> 16#0000_0000) AND (#Concatenadora <> 16#0000_0001) AND (#Concatenadora <> 16#0000_0002) AND (#Concatenadora <> 16#0000_0004) AND (#Concatenadora <> 16#0000_0008) AND (#Concatenadora <> 16#0000_0010) AND (#Concatenadora <> 16#0000_0020) AND (#Concatenadora <> 16#0000_0040) AND (#Concatenadora <> 16#0000_0080) AND (#Concatenadora <> 16#0000_0100) AND (#Concatenadora <> 16#0000_0200) AND (#Concatenadora <> 16#0000_0400) AND (#Concatenadora <> 16#0000_0800) AND (#Concatenadora <> 16#0000_1000) AND (#Concatenadora <> 16#0000_2000) AND (#Concatenadora <> 16#0000_4000) AND (#Concatenadora <> 16#0000_8000) AND (#Concatenadora <> 16#0001_0000) AND (#Concatenadora <> 16#0002_0000) AND (#Concatenadora <> 16#0004_0000) AND (#Concatenadora <> 16#0008_0000) AND (#Concatenadora <> 16#0010_0000) AND (#Concatenadora <> 16#0020_0000) AND (#Concatenadora <> 16#0040_0000) AND (#Concatenadora <> 16#0080_0000) AND (#Concatenadora <> 16#0100_0000) AND (#Concatenadora <> 16#0200_0000) AND (#Concatenadora <> 16#0400_0000) AND (#Concatenadora <> 16#0800_0000) AND (#Concatenadora <> 16#1000_0000) AND (#Concatenadora <> 16#2000_0000) AND (#Concatenadora <> 16#4000_0000) AND (#Concatenadora <> 16#8000_0000);
END_REGION

REGION Network 3: Estado 1
   RUNG wire#powerrail
      { S7_Templates := "SrcType := DWord" } EQ_Contact(in1 := #Prioritaria, in2 := 16#0000_0000)
      { S7_Templates := "SrcType := DWord" } EQ_Contact(in1 := #Concatenadora, in2 := 16#0000_0001)
      wire#w1
      I_Contact( #"Falla Prioritarias" )
      I_Contact( #"Error Concatenadoras" )
      { S7_GenerateENO := "TRUE" } Move(in := 16#0000_0001, out1 => #Estado)
   END_RUNG
   RUNG wire#powerrail
      { S7_Templates := "SrcType := DWord" } EQ_Contact(in1 := #Prioritaria, in2 := 16#0000_0001)
   END_RUNG wire#w1
   // the same network as SCL:
   IF (((#Prioritaria = 16#0000_0000) AND (#Concatenadora = 16#0000_0001)) OR (#Prioritaria = 16#0000_0001)) AND NOT #"Falla Prioritarias" AND NOT #"Error Concatenadoras" THEN
       #Estado := 16#0000_0001;
   END_IF;
END_REGION

REGION Network 4: Estado 2
   RUNG wire#powerrail
      { S7_Templates := "SrcType := DWord" } EQ_Contact(in1 := #Prioritaria, in2 := 16#0000_0000)
      { S7_Templates := "SrcType := DWord" } EQ_Contact(in1 := #Concatenadora, in2 := 16#0000_0002)
      wire#w1
      I_Contact( #"Falla Prioritarias" )
      I_Contact( #"Error Concatenadoras" )
      { S7_GenerateENO := "TRUE" } Move(in := 16#0000_0002, out1 => #Estado)
   END_RUNG
   RUNG wire#powerrail
      { S7_Templates := "SrcType := DWord" } EQ_Contact(in1 := #Prioritaria, in2 := 16#0000_0002)
   END_RUNG wire#w1
   // the same network as SCL:
   IF (((#Prioritaria = 16#0000_0000) AND (#Concatenadora = 16#0000_0002)) OR (#Prioritaria = 16#0000_0002)) AND NOT #"Falla Prioritarias" AND NOT #"Error Concatenadoras" THEN
       #Estado := 16#0000_0002;
   END_IF;
END_REGION

